screen "Dev_PID" 800x480, template "Settings"
   IOField "I/O field_8" at 170,11 size 171x26; FormatPattern ????????????????
      ProcessValue <- "PIDx_Name"
   Button "Button_1" at 165,265 size 112x32; TextOff 'DB 900 / DB 700'; Authorization "User administration"
      on Release: SetTag("PIDx", 900); SetTag("PIDx_Name", 'DB 900')
      Visibility <- "Support_DB_All_PIDs"
      Appearance <- "PIDx"
   Button "Button_4" at 165,305 size 112x32; TextOff 'DB 901 / DB 701'; Authorization "User administration"
      on Release: SetTag("PIDx", 901); SetTag("PIDx_Name", 'DB 901')
      Visibility <- "Support_DB_All_PIDs"
      Appearance <- "PIDx"
   Button "Button_17" at 165,345 size 112x32; TextOff 'DB 902 / DB 702'; Authorization "User administration"
      on Release: SetTag("PIDx", 902); SetTag("PIDx_Name", 'DB 902')
      Visibility <- "Support_DB_All_PIDs"
      Appearance <- "PIDx"
   Button "Button_6" at 165,385 size 112x32; TextOff 'DB 903 / DB 703'; Authorization "User administration"
      on Release: SetTag("PIDx", 903); SetTag("PIDx_Name", 'DB 903')
      Visibility <- "Support_DB_All_PIDs"
      Appearance <- "PIDx"
   Button "Button_15" at 443,265 size 112x32; TextOff 'DB 910 / DB 710'; Authorization "User administration"
      on Release: SetTag("PIDx", 910); SetTag("PIDx_Name", 'DB 910')
      Visibility <- "Support_DB_All_PIDs"
      Appearance <- "PIDx"
   Button "Button_18" at 443,305 size 112x32; TextOff 'DB 911 / DB 711'; Authorization "User administration"
      on Release: SetTag("PIDx", 911); SetTag("PIDx_Name", 'DB 911')
      Visibility <- "Support_DB_All_PIDs"
      Appearance <- "PIDx"
   Button "Button_23" at 443,345 size 112x32; TextOff 'DB 912 / DB 712'; Authorization "User administration"
      on Release: SetTag("PIDx", 912); SetTag("PIDx_Name", 'DB 912')
      Visibility <- "Support_DB_All_PIDs"
      Appearance <- "PIDx"
   Button "Button_24" at 443,385 size 112x32; TextOff 'DB 913 / DB 713'; Authorization "User administration"
      on Release: SetTag("PIDx", 913); SetTag("PIDx_Name", 'DB 913')
      Visibility <- "Support_DB_All_PIDs"
      Appearance <- "PIDx"
   Button "Button_25" at 443,425 size 112x32; TextOff 'DB 914 / DB 714'; Authorization "User administration"
      on Release: SetTag("PIDx", 914); SetTag("PIDx_Name", 'DB 914')
      Visibility <- "Support_DB_All_PIDs"
      Appearance <- "PIDx"
   Button "Button_26" at 583,344 size 112x32; TextOff 'DB 917 / DB 717'; Authorization "User administration"
      on Release: SetTag("PIDx", 917); SetTag("PIDx_Name", 'DB 917')
      Visibility <- "Support_DB_All_PIDs"
      Appearance <- "PIDx"
   Button "Button_29" at 583,384 size 112x32; TextOff 'DB 918 / DB 718'; Authorization "User administration"
      on Release: SetTag("PIDx", 918); SetTag("PIDx_Name", 'DB 918')
      Visibility <- "Support_DB_All_PIDs"
      Appearance <- "PIDx"
   Button "Button_31" at 583,264 size 112x32; TextOff 'DB 915 / DB 715'; Authorization "User administration"
      on Release: SetTag("PIDx", 915); SetTag("PIDx_Name", 'DB 915')
      Visibility <- "Support_DB_All_PIDs"
      Appearance <- "PIDx"
   Button "Button_32" at 583,304 size 112x32; TextOff 'DB 916 / DB 716'; Authorization "User administration"
      on Release: SetTag("PIDx", 916); SetTag("PIDx_Name", 'DB 916')
      Visibility <- "Support_DB_All_PIDs"
      Appearance <- "PIDx"
   Button "Button_33" at 165,425 size 112x32; TextOff 'DB 904 / DB 704'; Authorization "User administration"
      on Release: SetTag("PIDx", 904); SetTag("PIDx_Name", 'DB 904')
      Visibility <- "Support_DB_All_PIDs"
      Appearance <- "PIDx"
   Button "Button_34" at 583,424 size 112x32; TextOff 'DB 919 / DB 719'; Authorization "User administration"
      on Release: SetTag("PIDx", 919); SetTag("PIDx_Name", 'DB 919')
      Visibility <- "Support_DB_All_PIDs"
      Appearance <- "PIDx"
   Button "Button_35" at 304,265 size 112x32; TextOff 'DB 905 / DB 705'; Authorization "User administration"
      on Release: SetTag("PIDx", 905); SetTag("PIDx_Name", 'DB 905')
      Visibility <- "Support_DB_All_PIDs"
      Appearance <- "PIDx"
   Button "Button_36" at 304,305 size 112x32; TextOff 'DB 906 / DB 706'; Authorization "User administration"
      on Release: SetTag("PIDx", 906); SetTag("PIDx_Name", 'DB 906')
      Visibility <- "Support_DB_All_PIDs"
      Appearance <- "PIDx"
   Button "Button_37" at 304,345 size 112x32; TextOff 'DB 907 / DB 707'; Authorization "User administration"
      on Release: SetTag("PIDx", 907); SetTag("PIDx_Name", 'DB 907')
      Visibility <- "Support_DB_All_PIDs"
      Appearance <- "PIDx"
   Button "Button_38" at 304,385 size 112x32; TextOff 'DB 908 / DB 708'; Authorization "User administration"
      on Release: SetTag("PIDx", 908); SetTag("PIDx_Name", 'DB 908')
      Visibility <- "Support_DB_All_PIDs"
      Appearance <- "PIDx"
   Button "Button_39" at 304,425 size 112x32; TextOff 'DB 909 / DB 709'; Authorization "User administration"
      on Release: SetTag("PIDx", 909); SetTag("PIDx_Name", 'DB 909')
      Visibility <- "Support_DB_All_PIDs"
      Appearance <- "PIDx"
   Button "Button_7" at 251,41 size 90x22; TextOff 'Авто'; Authorization "Operate"; TextList "Hand"
      on Click: InvertBit("PID_x_CMD_Hand")
      Appearance <- "PID_x_CMD_Hand"
      ProcessValue <- "PID_x_CMD_Hand"
   Button "Button_8" at 251,107 size 90x22; TextOff 'Принудит. / Стоп'; Authorization "Operate"
      on Click: InvertBit("PID_x_CMD_Force")
      Appearance <- "PID_x_CMD_Force"
   Button "Button_13" at 251,74 size 90x22; TextOff 'Работа / Пуск'; Authorization "Operate"
      on Click: InvertBit("PID_x_CMD_Start_A")
      Appearance <- "PID_x_CMD_Start_A"
   Button "Button_19" at 251,140 size 90x22; TextOff 'Сброс аварий'; Authorization "Operate"
      on Click: SetBit("PID_x_CMD_Reset")
      Appearance <- "PID_x_CMD_Alarm"
   TextField "Text field_1" at 539,100 size 86x18; Text 'Мертвая зона:'
   IOField "I/O field_24" at 627,99 size 50x20; Authorization "User administration"; FormatPattern s99.99
      ProcessValue <- "PID_x_Settings_DeadBand"
   IOField "I/O field_9" at 627,121 size 50x20; Authorization "User administration"; FormatPattern 99.9
      ProcessValue <- "PID_x_C_SP"
   TextField "Text field_5" at 515,122 size 110x18; Text 'Частота вызова, с:'
   IOField "I/O field_10" at 377,29 size 55x20; Authorization "User administration"; FormatPattern s99.999
      ProcessValue <- "PID_x_Settings_SP_P"
   TextField "Text field_10" at 344,30 size 31x18; Text 'K'
   TextField "Text field_12" at 344,52 size 31x18; Text 'Ti'
   IOField "I/O field_12" at 377,50 size 55x20; Authorization "User administration"; FormatPattern 9999
      ProcessValue <- "PID_x_Settings_SP_Ti"
   IOField "I/O field_28" at 377,71 size 55x20; Authorization "User administration"; FormatPattern 9999
      ProcessValue <- "PID_x_Settings_SP_Td"
   TextField "Text field_6" at 345,72 size 31x18; Text 'Td'
   TextField "Text field_2" at 460,28 size 54x18; Text 'Уставка'
   IOField "I/O field_1" at 556,27 size 55x20; Authorization "User administration"; FormatPattern s9999.9
      ProcessValue <- "PID_x_Settings_Min_SP"
      Appearance <- "PID_x_Sys_Alm_SP_L"
   IOField "I/O field_2" at 620,27 size 55x20; Authorization "User administration"; FormatPattern s99999.9
      ProcessValue <- "PID_x_Settings_Max_SP"
      Appearance <- "PID_x_Sys_Alm_SP_H"
   TextField "Text field_4" at 572,8 size 31x18; Text 'от'
   TextField "Text field_7" at 635,8 size 31x18; Text 'до'
   TextField "Text field_8" at 460,52 size 50x18; Text 'Датчик'
   IOField "I/O field_3" at 556,51 size 55x20; Authorization "User administration"; FormatPattern s9999.9
      ProcessValue <- "PID_x_Settings_Min_in"
      Appearance <- "PID_x_Sys_Alm_In_L"
   IOField "I/O field_4" at 620,51 size 55x20; Authorization "User administration"; FormatPattern s99999.9
      ProcessValue <- "PID_x_Settings_Max_in"
      Appearance <- "PID_x_Sys_Alm_In_H"
   TextField "Text field_11" at 460,76 size 78x18; Text 'Выход ПИД'
   IOField "I/O field_7" at 556,75 size 55x20; Authorization "User administration"; FormatPattern s999.99
      ProcessValue <- "PID_x_Settings_Min_out"
   IOField "I/O field_5" at 620,75 size 55x20; Authorization "User administration"; FormatPattern s999.99
      ProcessValue <- "PID_x_Settings_Max_out"
   IOField "I/O field_6" at 433,99 size 55x20; Authorization "Developer"; FormatPattern 999.99
      ProcessValue <- "PID_x_x"
   TextField "Text field_3" at 345,100 size 86x18; Text 'Коэффициент'
   IOField "I/O field_11" at 171,54 size 78x25; Authorization "User administration"; FormatPattern s9999.9
      Appearance <- "PID_x_CMD_Hand"
      ProcessValue <- "PID_x_SP_M"
   TextField "Text field_22" at 177,36 size 68x18; Text 'Уставка / Показания:'
   IOField "I/O field_13" at 171,96 size 78x25; Authorization "User administration"; FormatPattern s9999.9
      ProcessValue <- "PID_x_Value"
   TextField "Text field_9" at 177,78 size 68x18; Text 'Датчик / Показания:'
   IOField "I/O field_14" at 171,139 size 78x25; Authorization "User administration"; FormatPattern s9999.9
      ProcessValue <- "PID_x_PID_Hand"
      Appearance <- "PID_x_CMD_Force"
   TextField "Text field_13" at 177,122 size 68x18; Text 'Выход ПИД / Показания:'
   TextField "Text field_14" at 345,122 size 104x18; Text 'Инверсия выхода'
   Button "Button_2" at 449,122 size 60x20; TextOff 'Text'; PictureList "ON_OFF"; Authorization "User administration"
      on Click: InvertBit("PID_x_CMD_Vector")
      ProcessValue <- "PID_x_CMD_Vector"
   IOField "I/O field_15" at 627,144 size 50x20; Authorization "User administration"; FormatPattern 99.9
      ProcessValue <- "PID_x_Settings_SP_Cycle"
   TextField "Text field_15" at 529,145 size 96x18; Text 'Время цикла, с:'
   IOField "I/O field_16" at 433,144 size 55x20; Authorization "Developer"; FormatPattern 9999999999
      ProcessValue <- "PID_x_Sys_Error_code"
   TextField "Text field_16" at 345,145 size 72x18; Text 'Код ошибки'
   SymbolicIOField "Symbolic I/O field_1" at 113,464 size 75x16; TextOn '1'; TextOff '0'; TextList "Hand"
      ProcessValue <- "PID_x_CMD_Hand"
   TextField "Text field_21" at 211,464 size 75x16; Text 'Уставка +1'
      Visibility <- "PID_x_CMD_Hand"
   TextField "Text field_17" at 311,464 size 75x16; Text 'Уставка -1'
      Visibility <- "PID_x_CMD_Hand"
   TextField "Text field_23" at 610,464 size 75x16; Text 'Сброс аварий'
   Softkey "Softkey_F7" at 0,0 size 0x0
      on KeyDown: SetBit("PID_x_CMD_Reset")
   Softkey "Softkey_F2" at 0,0 size 0x0
      on KeyDown: InvertBit("PID_x_CMD_Hand")
   Softkey "Softkey_F3" at 0,0 size 0x0
      on KeyDown: function_dd21b452("PID_x_SP_M", 1)
   Softkey "Softkey_F4" at 0,0 size 0x0
      on KeyDown: function_b9b71300("PID_x_SP_M", 1)
*)